// TIA Portal project "EMS" (V15.1)

(* hardware
DEVICE "HMI_SDC"  TP1500 Comfort
   slot 0: "HMI_SDC"  TP1500 Comfort  6AV2 124-0QC02-0AX0  15.0.0.0
   slot 1: "HMI_RT_2"  TP1500 Comfort  6AV2 124-0QC02-0AX0  15.0.0.0
   slot 5: "HMI_SDC._CP_2"  PROFINET Interface  15.0.0.0
      slot 1: "PROFINET Schnittstelle_1"  PROFINET Interface
         slot 1: "Port_1"  Port
         slot 2: "Port_2"  Port
   slot 6: "HMI_SDC._CP_1"  PROFINET Interface  15.0.0.0
      slot 1: "PROFINET Schnittstelle_GBit"  PROFINET Interface
         slot 1: "Port_1"  Port
   slot 7: "HMI_SDC.I/DP_CP_1"  MPI/DP Interface  15.0.0.0
DEVICE "SCALANCE W client"  SCALANCE W-Station
   slot 0: "SCALANCE W rack"  Rail
   slot 0: "_wlan"  SCALANCE W734-1 RJ45 US  6GK5 734-1FX00-0AB0  V6.2
DEVICE "S71500/ET200MP station_1"  S7-1500 station
   slot 0: "Rail_0"  Rack  6ES7 590-1***0-0AA0
   slot 1: "SDC_PLC"  CPU 1518-4 PN/DP  6ES7 518-4AP00-0AB0  V2.6
      slot 3: "CPU display_1"  6ES7591-1BA00-0AA0
   slot 2: "DI 16x24VDC BA_1"  DI 16x24VDC BA  6ES7 521-1BH10-0AA0  V1.0
   slot 3: "DQ 16x24VDC/0.5A BA_1"  DQ 16x24VDC/0.5A BA  6ES7 522-1BH10-0AA0  V1.0
DEVICE "ET 200SP station_2"  ET 200SP-Station
   slot 0: "Rack_0"  Rack  6ES5 710-8MAx1
   slot 1: "_PLC"  CPU 1512SP F-1 PN  6ES7 512-1SK01-0AB0  V2.1
   slot 2: "F-DI 8x24VDC HF_1"  F-DI 8x24VDC HF  6ES7 136-6BA00-0CA0  V1.0
      slot 1: "F-DI 8x24VDC HF_1"  F-DI 8x24VDC HF
   slot 3: "F-DQ 4x24VDC/2A PM HF_1"  F-DQ 4x24VDC/2A PM HF  6ES7 136-6DB00-0CA0  V1.0
      slot 1: "F-DQ 4x24VDC/2A PM HF_1"  F-DQ 4x24VDC/2A PM HF
   slot 4: "DI 16x24VDC ST_1"  DI 16x24VDC ST  6ES7 131-6BH00-0BA0  V1.1
      slot 1: "DI 16x24VDC ST_1"  DI 16x24VDC ST
   slot 5: "DQ 8x24VDC/0.5A ST_1"  DQ 8x24VDC/0.5A ST  6ES7 132-6BF01-0BA0  V0.0
      slot 1: "DQ 8x24VDC/0.5A ST_1"  DQ 8x24VDC/0.5A ST
   slot 6: "Server module_1"  Server module  6ES7 193-6PA00-0AA0  V1.1
      slot 1: "Server module_1"  Server module
   slot 127: "BA 2xRJ45"  BA 2xRJ45  6ES7 193-6AR00-0AA0  V0.0
      slot 32769: "Port_1"  6ES7 193-6AR00-0AA0
      slot 32770: "Port_2"  6ES7 193-6AR00-0AA0
DEVICE "GSD device_4"  GSD.Device.PN
   slot 0: "Rack"  Rack  V1.0
   slot 0: "_DRIVE"  SINAMICS G120D CU240D-2 PN(-F) V4.7  6SL3 544-0FB2x-1Fxx  V4.70
      slot 0: "SINAMICS G120D CU240D-2 PN(-F) V4.7"  SINAMICS G120D CU240D-2 PN(-F) V4.7
      slot 1: "PN-IO"  PN-IO
         slot 1: "Port 1"  Port 1
         slot 2: "Port 2"  Port 2
      slot 1: "Drive_1"  Drive
         slot 0: "Module Access Point"  Module Access Point
   slot 2: "SIEMENS telegram 352, PZD-6/6"  SIEMENS telegram 352, PZD-6/6
DEVICE "GSD device_1"  GSD.Device.PN
   slot 0: "Rack"  Rack  V1.0
   slot 0: "_ENCODER"  PCV-F200-B17-6011 Position Encoder  PXVxx-F200-B17-V1D-6011
      slot 0: "PCV-F200-B17-6011 Position Encoder"  PCV-F200-B17-6011 Position Encoder
      slot 1: "Interface"  Interface
         slot 1: "Port 1"  Port 1
         slot 2: "Port 2"  Port 2
      slot 1: "Configuration_1"  Configuration
         slot 0: "Configuration"  Configuration
   slot 2: "status_1"  status
      slot 0: "status"  status
   slot 3: "x position_1"  x position
      slot 0: "x position"  x position
   slot 4: "y position_1"  y position
      slot 0: "y position"  y position
DEVICE "GSD device_6"  GSD.Device.PN
   slot 0: "Rack"  Rack  V1.0
   slot 0: "_HMI"  IRD400  6ES7 292-0AA50-1AA0  R01.00.00
      slot 0: "IRD400"  IRD400
      slot 1: "PNIO"  PNIO
         slot 1: "Port 1"  Port 1
         slot 2: "Port 2"  Port 2
      slot 1: "IR Remote Control_1"  IR Remote Control
         slot 0: "IR Remote Control"  IR Remote Control
      slot 2: "Display and LED _1"  Display and LED 
         slot 0: "Display and LED"  Display and LED 
      slot 3: "DIO_1"  DIO
         slot 0: "DIO"  DIO
      slot 4: "IR-P2P_1"  IR-P2P
         slot 0: "IR-P2P"  IR-P2P
      slot 5: "Device Control_1"  Device Control
         slot 0: "Device Control"  Device Control
DEVICE "SCALANCE W access point"  SCALANCE W-Station
   slot 0: "SCALANCE W rack"  Rail
   slot 0: "WLAN_1"  SCALANCE W788-1 M12 US  6GK5 788-1GD00-0AB0  V6.2
DEVICE "GSD device_11"  GSD.Device.PN
   slot 0: "Rack"  Rack  V1.0
   slot 0: "plx32-pnd"  PLX32-EIP-PND  EPD2  1.02.002
      slot 0: "PLX32-EIP-PND"  PLX32-EIP-PND
      slot 1: "Interface1"  Interface1
         slot 1: "Port1"  Port1
   slot 1: "INPUT 512 Byte_1"  INPUT 512 Byte
      slot 0: "INPUT 512 Byte"  INPUT 512 Byte
   slot 2: "OUTPUT 512 Byte_1"  OUTPUT 512 Byte
      slot 0: "OUTPUT 512 Byte"  OUTPUT 512 Byte
   slot 3: "INPUT 256 Byte_3"  INPUT 256 Byte
      slot 0: "INPUT 256 Byte"  INPUT 256 Byte
   slot 4: "OUTPUT 256 Byte_3"  OUTPUT 256 Byte
      slot 0: "OUTPUT 256 Byte"  OUTPUT 256 Byte
   slot 5: "INPUT 256 Byte_2"  INPUT 256 Byte
      slot 0: "INPUT 256 Byte"  INPUT 256 Byte
   slot 6: "OUTPUT 256 Byte_2"  OUTPUT 256 Byte
      slot 0: "OUTPUT 256 Byte"  OUTPUT 256 Byte
   slot 7: "INPUT 256 Byte_1"  INPUT 256 Byte
      slot 0: "INPUT 256 Byte"  INPUT 256 Byte
   slot 8: "OUTPUT 256 Byte_1"  OUTPUT 256 Byte
      slot 0: "OUTPUT 256 Byte"  OUTPUT 256 Byte
*)

// ===== PLC "SDC_PLC"  CPU 1518-4 PN/DP =====

VAR_GLOBAL   // PLC tag table "Default tag table"
   "LinePLC1_RD_ready" AT %I4248.0 : Bool;
   "EMS_ProductionSpeedRef" AT %IW6130 : Word;
   "EMS_CarrierSpeedRef" AT %IW6126 : Word;
   "SDC_C2_OUT_W9" AT %QW468 : Word;
   "System_Byte" AT %MB1 : Byte;
   "FirstScan" AT %M1.0 : Bool;
   "DiagStatusUpdate" AT %M1.1 : Bool;
   "AlwaysTRUE" AT %M1.2 : Bool;
   "AlwaysFALSE" AT %M1.3 : Bool;
   "Clock_Byte" AT %MB0 : Byte;
   "Clock_10Hz" AT %M0.0 : Bool;
   "Clock_5Hz" AT %M0.1 : Bool;
   "Clock_2.5Hz" AT %M0.2 : Bool;
   "Clock_2Hz" AT %M0.3 : Bool;
   "Clock_1.25Hz" AT %M0.4 : Bool;
   "Clock_1Hz" AT %M0.5 : Bool;
   "Clock_0.625Hz" AT %M0.6 : Bool;
   "Clock_0.5Hz" AT %M0.7 : Bool;
   "tem" AT %M2.0 : Bool;
   "reset" AT %M2.1 : Bool;
   "ZoneCnt" AT %MW4 : Int;
   "Totalcar" AT %MW6 : Int;
   "Tag_3" AT %M2.2 : Bool;
   "carrierzone" AT %MW8 : Int;
   "Carriercnt" AT %MW10 : Int;
   "Carriercnt(1)" AT %MW12 : Int;
   "carrposn" AT %MW14 : Int;
   "IndexArraytemp" AT %MW20 : Int;
   "tempsort" AT %M2.4 : Bool;
   "tempenable2" AT %M2.5 : Bool;
   "tempenable3" AT %M2.6 : Bool;
   "tempenable4" AT %M2.7 : Bool;
   "tempenable5" AT %M3.0 : Bool;
   "tempenable7" AT %M3.1 : Bool;
   "tempblock" AT %M3.2 : Bool;
   "CarrierCounterGbl" AT %MW16 : Int;
   "temp" AT %M3.3 : Bool;
   "cARRIERTESTPOINT" AT %MW18 : Int;
   "cARRIERTESTPOINTBOOL" AT %M3.4 : Bool;
   "cARIERLOOPCOUNT" AT %MW22 : Int;
   "cARIERLOOPCOUNT2" AT %MW24 : Int;
   "tempcarrier27cmdfwd" AT %MW26 : Int;
   "tempcarrier27cmdfwd1" AT %M3.5 : Bool;
   "ZoneCounterGbl" AT %MW28 : Int;
   "IndiconTempDebugON" AT %M3.6 : Bool;
   "HMI_EMS_Nr" AT %MW30 : Int;
   "HMI_EMS_Nr_Calc1" AT %MW32 : Int;
   "HMI_EMS_Nr_Calc2" AT %MW34 : Int;
   "HMI_EMS_Nr__Flt_Out" AT %MW36 : Int;
   "HMI_EMS_Nr__Warn_Out" AT %MW38 : Int;
   "TrafficCopZoneArrayPosCounter" AT %MW40 : Int;
   "SectionComment" AT %M42.0 : Bool;
   "DuplicateCarrierfound" AT %M42.1 : Bool;
   "FaultReset" AT %M42.2 : Bool;
   "DuplicateCarrierNumber" AT %MW44 : Word;
   "CarrierNumberLoop" AT %MW46 : Int;
   "Zone5_ClearToEnter" AT %M42.3 : Bool;
   "PrevCarrierInTransitMem" AT %M42.4 : Bool;
   "SecondDuplicateCarrierPosition" AT %MW50 : Word;
   "FirstDuplicateCarrierPosition" AT %MW48 : Word;
   "EMS_Fault_Reset" AT %M42.5 : Bool;
   "TCCarrierCounterGbl" AT %MW100 : Int;
   "FC206CarrierLoop" AT %MW52 : Int;
   "FC206PositionLoop" AT %MW54 : Int;
   "CARRIER01_POSITION_SDC_OUT" AT %ID402 : DWord;
   "Temp_Int" AT %MW56 : Int;
   "CARRIER #01   1 STATUS [0].5" AT %M80.5 : Bool;
   "CARRIER #01   CURRENT" AT %MW72 : Int;
   "CARRIER #01   G120D CONTROL WORD.0" AT %M74.0 : Bool;
   "CARRIER #01   G120D CONTROL WORD.1" AT %M74.1 : Bool;
   "CARRIER #01   G120D CONTROL WORD.10" AT %M75.2 : Bool;
   "CARRIER #01   G120D CONTROL WORD.11" AT %M75.3 : Bool;
   "CARRIER #01   G120D CONTROL WORD.12" AT %M75.4 : Bool;
   "CARRIER #01   G120D CONTROL WORD.13" AT %M75.5 : Bool;
   "CARRIER #01   G120D CONTROL WORD.14" AT %M75.6 : Bool;
   "CARRIER #01   G120D CONTROL WORD.15" AT %M75.7 : Bool;
   "CARRIER #01   G120D CONTROL WORD.2" AT %M74.2 : Bool;
   "CARRIER #01   G120D CONTROL WORD.3" AT %M74.3 : Bool;
   "CARRIER #01   G120D CONTROL WORD.4" AT %M74.4 : Bool;
   "CARRIER #01   G120D CONTROL WORD.5" AT %M74.5 : Bool;
   "CARRIER #01   G120D CONTROL WORD.6" AT %M74.6 : Bool;
   "CARRIER #01   G120D CONTROL WORD.7" AT %M74.7 : Bool;
   "CARRIER #01   G120D CONTROL WORD.8" AT %M75.0 : Bool;
   "CARRIER #01   G120D CONTROL WORD.9" AT %M75.1 : Bool;
   "CARRIER #01   G120D STATUS WORD.0" AT %M76.0 : Bool;
   "CARRIER #01   G120D STATUS WORD.1" AT %M76.1 : Bool;
   "CARRIER #01   G120D STATUS WORD.10" AT %M77.2 : Bool;
   "CARRIER #01   G120D STATUS WORD.11" AT %M77.3 : Bool;
   "CARRIER #01   G120D STATUS WORD.12" AT %M77.4 : Bool;
   "CARRIER #01   G120D STATUS WORD.13" AT %M77.5 : Bool;
   "CARRIER #01   G120D STATUS WORD.14" AT %M77.6 : Bool;
   "CARRIER #01   G120D STATUS WORD.15" AT %M77.7 : Bool;
   "CARRIER #01   G120D STATUS WORD.2" AT %M76.2 : Bool;
   "CARRIER #01   G120D STATUS WORD.3" AT %M76.3 : Bool;
   "CARRIER #01   G120D STATUS WORD.4" AT %M76.4 : Bool;
   "CARRIER #01   G120D STATUS WORD.5" AT %M76.5 : Bool;
   "CARRIER #01   G120D STATUS WORD.6" AT %M76.6 : Bool;
   "CARRIER #01   G120D STATUS WORD.7" AT %M76.7 : Bool;
   "CARRIER #01   G120D STATUS WORD.8" AT %M77.0 : Bool;
   "CARRIER #01   G120D STATUS WORD.9" AT %M77.1 : Bool;
   "CARRIER #01   POSITION" AT %MW78 : Int;
   "CARRIER #01 480VPowerOn_MDCB1" AT %M80.0 : Bool;
   "CARRIER #01 CrashDetectSW" AT %M80.1 : Bool;
   "CARRIER #01 DCsupplyOnPSCB2" AT %M80.2 : Bool;
   "CARRIER #01 FaultLight_LH" AT %M80.3 : Bool;
   "CARRIER #01 FaultLight_RH" AT %M80.4 : Bool;
   "CARRIER #01 PB1_ProdHoldLH" AT %M80.6 : Bool;
   "CARRIER #01 PB2_ResetLH" AT %M80.7 : Bool;
   "CARRIER #01 PB3_ProdHoldRH" AT %M81.0 : Bool;
   "CARRIER #01 PB4_ResetRH" AT %M81.1 : Bool;
   "CARRIER #01 RunLight_LH" AT %M81.2 : Bool;
   "CARRIER #01 RunLight_RH" AT %M81.3 : Bool;
   "CARRIER #01 SitopSelectStatus" AT %M81.4 : Bool;
   "CARRIER #01 SpareInput(2_1)" AT %M81.5 : Bool;
   "CARRIER #01 SpareInput(2_2)" AT %M81.6 : Bool;
   "CARRIER #01 SpareInput(2_3)" AT %M81.7 : Bool;
   "CARRIER #01 SpareInput(2_4)" AT %M82.0 : Bool;
   "CARRIER #01 SpareInput(2_5)" AT %M82.1 : Bool;
   "CARRIER #01 SpareInput(2_6)" AT %M82.2 : Bool;
   "CARRIER #01 SpareInput(2_7)" AT %M82.3 : Bool;
   "CARRIER #01 SpareInput(4_1)" AT %M82.4 : Bool;
   "CARRIER #01 SpareInput(4_14)" AT %M82.5 : Bool;
   "CARRIER #01 SpareInput(4_15)" AT %M82.6 : Bool;
   "CARRIER #01 SpareInput(4_16)" AT %M82.7 : Bool;
   "CARRIER #01 SpareInput(4_17)" AT %M83.0 : Bool;
   "CARRIER #01 SpareInput(4_2)" AT %M83.1 : Bool;
   "CARRIER #01 SpareInput(4_5)" AT %M83.2 : Bool;
   "CARRIER #01 SpareInput(4_6)" AT %M83.3 : Bool;
   "CARRIER #01 SpareInput(4_7)" AT %M83.4 : Bool;
   "CARRIER #01 SpareOutput(5_5)" AT %M83.5 : Bool;
   "CARRIER #01 SpareOutput(5_6)" AT %M83.6 : Bool;
   "CARRIER #01 SpareOutput(5_7)" AT %M83.7 : Bool;
   "CARRIER #01 SpareSafetyOutput(3_1)" AT %M84.0 : Bool;
   "CARRIER #01 SpareSafetyOutput(3_2)" AT %M84.1 : Bool;
   "CARRIER #01 SpareSafetyOutput(3_3)" AT %M84.2 : Bool;
   "CARRIER #01 SpareSafetyOutput(3_4)" AT %M84.3 : Bool;
   "CARRIER #01 SpareSafetyOutput(3_5)" AT %M84.4 : Bool;
   "CARRIER #01 SpareSafetyOutput(3_6)" AT %M84.5 : Bool;
   "CARRIER #01 SpareSafetyOutput(3_7)" AT %M84.6 : Bool;
   "Carrier #01_ At Command Position" AT %M84.7 : Bool;
   "Carrier #01_ Carrier in zone" AT %MW86 : Int;
   "Carrier #01_ Next carrier number" AT %MW88 : Int;
   "Carrier 1  Drive Status" AT %I412.1 : Bool;
   "Carrier 1 HMI Status" AT %I412.2 : Bool;
   "Carrier 1 PnF Encoder Status" AT %I412.0 : Bool;
   "Carrier 1 Profinet Fault" AT %I410.7 : Bool;
   "Carrier 2  Drive Status" AT %I432.1 : Bool;
   "Carrier 2 HMI Status" AT %I432.2 : Bool;
   "Carrier 2 PnF Encoder Status" AT %I432.0 : Bool;
   "Carrier 2 Profinet Fault" AT %I430.7 : Bool;
   "Carrier 3  Drive Status" AT %I452.1 : Bool;
   "Carrier 3 HMI Status" AT %I452.2 : Bool;
   "Carrier 3 PnF Encoder Status" AT %I452.0 : Bool;
   "Carrier 4  Drive Status" AT %I472.1 : Bool;
   "Carrier 4 HMI Status" AT %I472.2 : Bool;
   "Carrier 4 PnF Encoder Status" AT %I472.0 : Bool;
   "Carrier 4 Profinet Fault" AT %I470.7 : Bool;
   "Carrier_Index_HMI" AT %MW70 : Int;
   "HMI_Zone_Nr" AT %MW102 : Int;
END_VAR

VAR_GLOBAL CONSTANT   // PLC tag table "UserDiag_Constants"
   "USERDIAG_IOSYSTEM_1" : Int := 1;   // Index for first IO-System/DP-Mastersystem
   "USERDIAG_IOSYSTEM_2" : Int := 2;   // Index for second IO-System/DP-Mastersystem
   "USERDIAG_DEVICES_PER_SCREEN_UPPER_LIM" : Int := 128;   // Upper limit of devices per HMI screen
   "USERDIAG_SLOTS_PER_SCREEN_UPPER_LIM" : Int := 31;   // Upper limit of slots per HMI screen
   "USERDIAG_SLOTS_PER_DEVICE_UPPER_LIM" : Int := 31;   // max number of modules per device
   "USERDIAG_DEVICES_PER_IO_SYSTEM_UPPER_LIM" : Int := 128;   // Upper limit of devices/slaves per IO-System/DP-Mastersystem
   "USERDIAG_SLOTS_PER_PLC_UPPER_LIM" : Int := 31;   // max number of local modules
   "USERDIAG_IO_SYSTEMS_UPPER_LIM" : Int := 2;   // Upper limit of IO-Systems/DP-Mastersystems
   "USERDIAG_IOSYSTEM_3" : Int := 3;   // Index for third IO-System/DP-Mastersystem
END_VAR

VAR_GLOBAL   // PLC tag table "SDC_AB_TagTable"
   "SDC_EMS01_CARRIER1_Spare0" AT %Q6768.0 : Bool;
   "SDC_EMS01_CARRIER1_DriveTripped" AT %Q6768.1 : Bool;
   "SDC_EMS01_CARRIER1_Spare2" AT %Q6768.2 : Bool;
   "SDC_EMS01_CARRIER1_PositioningComplete" AT %Q6768.3 : Bool;
   "SDC_EMS01_CARRIER1_RunStopPressed" AT %Q6768.4 : Bool;
   "SDC_EMS01_CARRIER1_Moving" AT %Q6768.5 : Bool;
   "SDC_EMS01_CARRIER1_Faulted" AT %Q6768.6 : Bool;
   "SDC_EMS01_CARRIER1_InAuto" AT %Q6768.7 : Bool;
   "SDC_EMS01_CARRIER2_Spare0" AT %Q6769.0 : Bool;
   "SDC_EMS01_CARRIER2_DriveTripped" AT %Q6769.1 : Bool;
   "SDC_EMS01_CARRIER2_Spare2" AT %Q6769.2 : Bool;
   "SDC_EMS01_CARRIER2_PositioningComplete" AT %Q6769.3 : Bool;
   "SDC_EMS01_CARRIER2_RunStopPressed" AT %Q6769.4 : Bool;
   "SDC_EMS01_CARRIER2_Moving" AT %Q6769.5 : Bool;
   "SDC_EMS01_CARRIER2_Faulted" AT %Q6769.6 : Bool;
   "SDC_EMS01_CARRIER2_InAuto" AT %Q6769.7 : Bool;
   "SDC_EMS01_CARRIER3_Spare0" AT %Q6770.0 : Bool;
   "SDC_EMS01_CARRIER3_DriveTripped" AT %Q6770.1 : Bool;
   "SDC_EMS01_CARRIER3_Spare2" AT %Q6770.2 : Bool;
   "SDC_EMS01_CARRIER3_PositioningComplete" AT %Q6770.3 : Bool;
   "SDC_EMS01_CARRIER3_RunStopPressed" AT %Q6770.4 : Bool;
   "SDC_EMS01_CARRIER3_Moving" AT %Q6770.5 : Bool;
   "SDC_EMS01_CARRIER3_Faulted" AT %Q6770.6 : Bool;
   "SDC_EMS01_CARRIER3_InAuto" AT %Q6770.7 : Bool;
   "SDC_EMS01_CARRIER4_Spare0" AT %Q6771.0 : Bool;
   "SDC_EMS01_CARRIER4_DriveTripped" AT %Q6771.1 : Bool;
   "SDC_EMS01_CARRIER4_Spare2" AT %Q6771.2 : Bool;
   "SDC_EMS01_CARRIER4_PositioningComplete" AT %Q6771.3 : Bool;
   "SDC_EMS01_CARRIER4_RunStopPressed" AT %Q6771.4 : Bool;
   "SDC_EMS01_CARRIER4_Moving" AT %Q6771.5 : Bool;
   "SDC_EMS01_CARRIER4_Faulted" AT %Q6771.6 : Bool;
   "SDC_EMS01_CARRIER4_InAuto" AT %Q6771.7 : Bool;
   "SDC_EMS01_CARRIER5_Spare0" AT %Q6772.0 : Bool;
   "SDC_EMS01_CARRIER5_DriveTripped" AT %Q6772.1 : Bool;
   "SDC_EMS01_CARRIER5_Spare2" AT %Q6772.2 : Bool;
   "SDC_EMS01_CARRIER5_PositioningComplete" AT %Q6772.3 : Bool;
   "SDC_EMS01_CARRIER5_RunStopPressed" AT %Q6772.4 : Bool;
   "SDC_EMS01_CARRIER5_Moving" AT %Q6772.5 : Bool;
   "SDC_EMS01_CARRIER5_Faulted" AT %Q6772.6 : Bool;
   "SDC_EMS01_CARRIER5_InAuto" AT %Q6772.7 : Bool;
   "SDC_EMS01_CARRIER6_Spare0" AT %Q6773.0 : Bool;
   "SDC_EMS01_CARRIER6_DriveTripped" AT %Q6773.1 : Bool;
   "SDC_EMS01_CARRIER6_Spare2" AT %Q6773.2 : Bool;
   "SDC_EMS01_CARRIER6_PositioningComplete" AT %Q6773.3 : Bool;
   "SDC_EMS01_CARRIER6_RunStopPressed" AT %Q6773.4 : Bool;
   "SDC_EMS01_CARRIER6_Moving" AT %Q6773.5 : Bool;
   "SDC_EMS01_CARRIER6_Faulted" AT %Q6773.6 : Bool;
   "SDC_EMS01_CARRIER6_InAuto" AT %Q6773.7 : Bool;
   "SDC_EMS01_CARRIER7_Spare0" AT %Q6774.0 : Bool;
   "SDC_EMS01_CARRIER7_DriveTripped" AT %Q6774.1 : Bool;
   "SDC_EMS01_CARRIER7_Spare2" AT %Q6774.2 : Bool;
   "SDC_EMS01_CARRIER7_PositioningComplete" AT %Q6774.3 : Bool;
   "SDC_EMS01_CARRIER7_RunStopPressed" AT %Q6774.4 : Bool;
   "SDC_EMS01_CARRIER7_Moving" AT %Q6774.5 : Bool;
   "SDC_EMS01_CARRIER7_Faulted" AT %Q6774.6 : Bool;
   "SDC_EMS01_CARRIER7_InAuto" AT %Q6774.7 : Bool;
   "SDC_EMS01_CARRIER8_Spare0" AT %Q6775.0 : Bool;
   "SDC_EMS01_CARRIER8_DriveTripped" AT %Q6775.1 : Bool;
   "SDC_EMS01_CARRIER8_Spare2" AT %Q6775.2 : Bool;
   "SDC_EMS01_CARRIER8_PositioningComplete" AT %Q6775.3 : Bool;
   "SDC_EMS01_CARRIER8_RunStopPressed" AT %Q6775.4 : Bool;
   "SDC_EMS01_CARRIER8_Moving" AT %Q6775.5 : Bool;
   "SDC_EMS01_CARRIER8_Faulted" AT %Q6775.6 : Bool;
   "SDC_EMS01_CARRIER8_InAuto" AT %Q6775.7 : Bool;
   "SDC_EMS01_CARRIER9_Spare0" AT %Q6776.0 : Bool;
   "SDC_EMS01_CARRIER9_DriveTripped" AT %Q6776.1 : Bool;
   "SDC_EMS01_CARRIER9_Spare2" AT %Q6776.2 : Bool;
   "SDC_EMS01_CARRIER9_PositioningComplete" AT %Q6776.3 : Bool;
   "SDC_EMS01_CARRIER9_RunStopPressed" AT %Q6776.4 : Bool;
   "SDC_EMS01_CARRIER9_Moving" AT %Q6776.5 : Bool;
   "SDC_EMS01_CARRIER9_Faulted" AT %Q6776.6 : Bool;
   "SDC_EMS01_CARRIER9_InAuto" AT %Q6776.7 : Bool;
   "SDC_EMS01_CARRIER10_Spare0" AT %Q6777.0 : Bool;
   "SDC_EMS01_CARRIER10_DriveTripped" AT %Q6777.1 : Bool;
   "SDC_EMS01_CARRIER10_Spare2" AT %Q6777.2 : Bool;
   "SDC_EMS01_CARRIER10_PositioningComplete" AT %Q6777.3 : Bool;
   "SDC_EMS01_CARRIER10_RunStopPressed" AT %Q6777.4 : Bool;
   "SDC_EMS01_CARRIER10_Moving" AT %Q6777.5 : Bool;
   "SDC_EMS01_CARRIER10_Faulted" AT %Q6777.6 : Bool;
   "SDC_EMS01_CARRIER10_InAuto" AT %Q6777.7 : Bool;
   "SDC_EMS01_CARRIER11_Spare0" AT %Q6778.0 : Bool;
   "SDC_EMS01_CARRIER11_DriveTripped" AT %Q6778.1 : Bool;
   "SDC_EMS01_CARRIER11_Spare2" AT %Q6778.2 : Bool;
   "SDC_EMS01_CARRIER11_PositioningComplete" AT %Q6778.3 : Bool;
   "SDC_EMS01_CARRIER11_RunStopPressed" AT %Q6778.4 : Bool;
   "SDC_EMS01_CARRIER11_Moving" AT %Q6778.5 : Bool;
   "SDC_EMS01_CARRIER11_Faulted" AT %Q6778.6 : Bool;
   "SDC_EMS01_CARRIER11_InAuto" AT %Q6778.7 : Bool;
   "SDC_EMS01_CARRIER12_Spare0" AT %Q6779.0 : Bool;
   "SDC_EMS01_CARRIER12_DriveTripped" AT %Q6779.1 : Bool;
   "SDC_EMS01_CARRIER12_Spare2" AT %Q6779.2 : Bool;
   "SDC_EMS01_CARRIER12_PositioningComplete" AT %Q6779.3 : Bool;
   "SDC_EMS01_CARRIER12_RunStopPressed" AT %Q6779.4 : Bool;
   "SDC_EMS01_CARRIER12_Moving" AT %Q6779.5 : Bool;
   "SDC_EMS01_CARRIER12_Faulted" AT %Q6779.6 : Bool;
   "SDC_EMS01_CARRIER12_InAuto" AT %Q6779.7 : Bool;
   "SDC_EMS01_CARRIER13_Spare0" AT %Q6780.0 : Bool;
   "SDC_EMS01_CARRIER13_DriveTripped" AT %Q6780.1 : Bool;
   "SDC_EMS01_CARRIER13_Spare2" AT %Q6780.2 : Bool;
   "SDC_EMS01_CARRIER13_PositioningComplete" AT %Q6780.3 : Bool;
   "SDC_EMS01_CARRIER13_RunStopPressed" AT %Q6780.4 : Bool;
   "SDC_EMS01_CARRIER13_Moving" AT %Q6780.5 : Bool;
   "SDC_EMS01_CARRIER13_Faulted" AT %Q6780.6 : Bool;
   "SDC_EMS01_CARRIER13_InAuto" AT %Q6780.7 : Bool;
   "SDC_EMS01_CARRIER14_Spare0" AT %Q6781.0 : Bool;
   "SDC_EMS01_CARRIER14_DriveTripped" AT %Q6781.1 : Bool;
   "SDC_EMS01_CARRIER14_Spare2" AT %Q6781.2 : Bool;
   "SDC_EMS01_CARRIER14_PositioningComplete" AT %Q6781.3 : Bool;
   "SDC_EMS01_CARRIER14_RunStopPressed" AT %Q6781.4 : Bool;
   "SDC_EMS01_CARRIER14_Moving" AT %Q6781.5 : Bool;
   "SDC_EMS01_CARRIER14_Faulted" AT %Q6781.6 : Bool;
   "SDC_EMS01_CARRIER14_InAuto" AT %Q6781.7 : Bool;
   "SDC_EMS01_CARRIER15_Spare0" AT %Q6782.0 : Bool;
   "SDC_EMS01_CARRIER15_DriveTripped" AT %Q6782.1 : Bool;
   "SDC_EMS01_CARRIER15_Spare2" AT %Q6782.2 : Bool;
   "SDC_EMS01_CARRIER15_PositioningComplete" AT %Q6782.3 : Bool;
   "SDC_EMS01_CARRIER15_RunStopPressed" AT %Q6782.4 : Bool;
   "SDC_EMS01_CARRIER15_Moving" AT %Q6782.5 : Bool;
   "SDC_EMS01_CARRIER15_Faulted" AT %Q6782.6 : Bool;
   "SDC_EMS01_CARRIER15_InAuto" AT %Q6782.7 : Bool;
   "SDC_EMS01_CARRIER16_Spare0" AT %Q6783.0 : Bool;
   "SDC_EMS01_CARRIER16_DriveTripped" AT %Q6783.1 : Bool;
   "SDC_EMS01_CARRIER16_Spare2" AT %Q6783.2 : Bool;
   "SDC_EMS01_CARRIER16_PositioningComplete" AT %Q6783.3 : Bool;
   "SDC_EMS01_CARRIER16_RunStopPressed" AT %Q6783.4 : Bool;
   "SDC_EMS01_CARRIER16_Moving" AT %Q6783.5 : Bool;
   "SDC_EMS01_CARRIER16_Faulted" AT %Q6783.6 : Bool;
   "SDC_EMS01_CARRIER16_InAuto" AT %Q6783.7 : Bool;
   "SDC_EMS01_CARRIER17_Spare0" AT %Q6784.0 : Bool;
   "SDC_EMS01_CARRIER17_DriveTripped" AT %Q6784.1 : Bool;
   "SDC_EMS01_CARRIER17_Spare2" AT %Q6784.2 : Bool;
   "SDC_EMS01_CARRIER17_PositioningComplete" AT %Q6784.3 : Bool;
   "SDC_EMS01_CARRIER17_RunStopPressed" AT %Q6784.4 : Bool;
   "SDC_EMS01_CARRIER17_Moving" AT %Q6784.5 : Bool;
   "SDC_EMS01_CARRIER17_Faulted" AT %Q6784.6 : Bool;
   "SDC_EMS01_CARRIER17_InAuto" AT %Q6784.7 : Bool;
   "SDC_EMS01_CARRIER18_Spare0" AT %Q6785.0 : Bool;
   "SDC_EMS01_CARRIER18_DriveTripped" AT %Q6785.1 : Bool;
   "SDC_EMS01_CARRIER18_Spare2" AT %Q6785.2 : Bool;
   "SDC_EMS01_CARRIER18_PositioningComplete" AT %Q6785.3 : Bool;
   "SDC_EMS01_CARRIER18_RunStopPressed" AT %Q6785.4 : Bool;
   "SDC_EMS01_CARRIER18_Moving" AT %Q6785.5 : Bool;
   "SDC_EMS01_CARRIER18_Faulted" AT %Q6785.6 : Bool;
   "SDC_EMS01_CARRIER18_InAuto" AT %Q6785.7 : Bool;
   "SDC_EMS01_CARRIER19_Spare0" AT %Q6786.0 : Bool;
   "SDC_EMS01_CARRIER19_DriveTripped" AT %Q6786.1 : Bool;
   "SDC_EMS01_CARRIER19_Spare2" AT %Q6786.2 : Bool;
   "SDC_EMS01_CARRIER19_PositioningComplete" AT %Q6786.3 : Bool;
   "SDC_EMS01_CARRIER19_RunStopPressed" AT %Q6786.4 : Bool;
   "SDC_EMS01_CARRIER19_Moving" AT %Q6786.5 : Bool;
   "SDC_EMS01_CARRIER19_Faulted" AT %Q6786.6 : Bool;
   "SDC_EMS01_CARRIER19_InAuto" AT %Q6786.7 : Bool;
   "SDC_EMS01_CARRIER20_Spare0" AT %Q6787.0 : Bool;
   "SDC_EMS01_CARRIER20_DriveTripped" AT %Q6787.1 : Bool;
   "SDC_EMS01_CARRIER20_Spare2" AT %Q6787.2 : Bool;
   "SDC_EMS01_CARRIER20_PositioningComplete" AT %Q6787.3 : Bool;
   "SDC_EMS01_CARRIER20_RunStopPressed" AT %Q6787.4 : Bool;
   "SDC_EMS01_CARRIER20_Moving" AT %Q6787.5 : Bool;
   "SDC_EMS01_CARRIER20_Faulted" AT %Q6787.6 : Bool;
   "SDC_EMS01_CARRIER20_InAuto" AT %Q6787.7 : Bool;
   "SDC_EMS01_CARRIER21_Spare0" AT %Q6788.0 : Bool;
   "SDC_EMS01_CARRIER21_DriveTripped" AT %Q6788.1 : Bool;
   "SDC_EMS01_CARRIER21_Spare2" AT %Q6788.2 : Bool;
   "SDC_EMS01_CARRIER21_PositioningComplete" AT %Q6788.3 : Bool;
   "SDC_EMS01_CARRIER21_RunStopPressed" AT %Q6788.4 : Bool;
   "SDC_EMS01_CARRIER21_Moving" AT %Q6788.5 : Bool;
   "SDC_EMS01_CARRIER21_Faulted" AT %Q6788.6 : Bool;
   "SDC_EMS01_CARRIER21_InAuto" AT %Q6788.7 : Bool;
   "SDC_EMS01_CARRIER22_Spare0" AT %Q6789.0 : Bool;
   "SDC_EMS01_CARRIER22_DriveTripped" AT %Q6789.1 : Bool;
   "SDC_EMS01_CARRIER22_Spare2" AT %Q6789.2 : Bool;
   "SDC_EMS01_CARRIER22_PositioningComplete" AT %Q6789.3 : Bool;
   "SDC_EMS01_CARRIER22_RunStopPressed" AT %Q6789.4 : Bool;
   "SDC_EMS01_CARRIER22_Moving" AT %Q6789.5 : Bool;
   "SDC_EMS01_CARRIER22_Faulted" AT %Q6789.6 : Bool;
   "SDC_EMS01_CARRIER22_InAuto" AT %Q6789.7 : Bool;
   "SDC_EMS01_CARRIER23_Spare0" AT %Q6790.0 : Bool;
   "SDC_EMS01_CARRIER23_DriveTripped" AT %Q6790.1 : Bool;
   "SDC_EMS01_CARRIER23_Spare2" AT %Q6790.2 : Bool;
   "SDC_EMS01_CARRIER23_PositioningComplete" AT %Q6790.3 : Bool;
   "SDC_EMS01_CARRIER23_RunStopPressed" AT %Q6790.4 : Bool;
   "SDC_EMS01_CARRIER23_Moving" AT %Q6790.5 : Bool;
   "SDC_EMS01_CARRIER23_Faulted" AT %Q6790.6 : Bool;
   "SDC_EMS01_CARRIER23_InAuto" AT %Q6790.7 : Bool;
   "SDC_EMS01_CARRIER24_Spare0" AT %Q6791.0 : Bool;
   "SDC_EMS01_CARRIER24_DriveTripped" AT %Q6791.1 : Bool;
   "SDC_EMS01_CARRIER24_Spare2" AT %Q6791.2 : Bool;
   "SDC_EMS01_CARRIER24_PositioningComplete" AT %Q6791.3 : Bool;
   "SDC_EMS01_CARRIER24_RunStopPressed" AT %Q6791.4 : Bool;
   "SDC_EMS01_CARRIER24_Moving" AT %Q6791.5 : Bool;
   "SDC_EMS01_CARRIER24_Faulted" AT %Q6791.6 : Bool;
   "SDC_EMS01_CARRIER24_InAuto" AT %Q6791.7 : Bool;
   "SDC_EMS01_CARRIER25_Spare0" AT %Q6792.0 : Bool;
   "SDC_EMS01_CARRIER25_DriveTripped" AT %Q6792.1 : Bool;
   "SDC_EMS01_CARRIER25_Spare2" AT %Q6792.2 : Bool;
   "SDC_EMS01_CARRIER25_PositioningComplete" AT %Q6792.3 : Bool;
   "SDC_EMS01_CARRIER25_RunStopPressed" AT %Q6792.4 : Bool;
   "SDC_EMS01_CARRIER25_Moving" AT %Q6792.5 : Bool;
   "SDC_EMS01_CARRIER25_Faulted" AT %Q6792.6 : Bool;
   "SDC_EMS01_CARRIER25_InAuto" AT %Q6792.7 : Bool;
   "SDC_EMS01_CARRIER26_Spare0" AT %Q6793.0 : Bool;
   "SDC_EMS01_CARRIER26_DriveTripped" AT %Q6793.1 : Bool;
   "SDC_EMS01_CARRIER26_Spare2" AT %Q6793.2 : Bool;
   "SDC_EMS01_CARRIER26_PositioningComplete" AT %Q6793.3 : Bool;
   "SDC_EMS01_CARRIER26_RunStopPressed" AT %Q6793.4 : Bool;
   "SDC_EMS01_CARRIER26_Moving" AT %Q6793.5 : Bool;
   "SDC_EMS01_CARRIER26_Faulted" AT %Q6793.6 : Bool;
   "SDC_EMS01_CARRIER26_InAuto" AT %Q6793.7 : Bool;
   "SDC_EMS01_CARRIER27_Spare0" AT %Q6794.0 : Bool;
   "SDC_EMS01_CARRIER27_DriveTripped" AT %Q6794.1 : Bool;
   "SDC_EMS01_CARRIER27_Spare2" AT %Q6794.2 : Bool;
   "SDC_EMS01_CARRIER27_PositioningComplete" AT %Q6794.3 : Bool;
   "SDC_EMS01_CARRIER27_RunStopPressed" AT %Q6794.4 : Bool;
   "SDC_EMS01_CARRIER27_Moving" AT %Q6794.5 : Bool;
   "SDC_EMS01_CARRIER27_Faulted" AT %Q6794.6 : Bool;
   "SDC_EMS01_CARRIER27_InAuto" AT %Q6794.7 : Bool;
   "SDC_EMS01_CARRIER28_Spare0" AT %Q6795.0 : Bool;
   "SDC_EMS01_CARRIER28_DriveTripped" AT %Q6795.1 : Bool;
   "SDC_EMS01_CARRIER28_Spare2" AT %Q6795.2 : Bool;
   "SDC_EMS01_CARRIER28_PositioningComplete" AT %Q6795.3 : Bool;
   "SDC_EMS01_CARRIER28_RunStopPressed" AT %Q6795.4 : Bool;
   "SDC_EMS01_CARRIER28_Moving" AT %Q6795.5 : Bool;
   "SDC_EMS01_CARRIER28_Faulted" AT %Q6795.6 : Bool;
   "SDC_EMS01_CARRIER28_InAuto" AT %Q6795.7 : Bool;
   "SDC_EMS01_CARRIER29_Spare0" AT %Q6796.0 : Bool;
   "SDC_EMS01_CARRIER29_DriveTripped" AT %Q6796.1 : Bool;
   "SDC_EMS01_CARRIER29_Spare2" AT %Q6796.2 : Bool;
   "SDC_EMS01_CARRIER29_PositioningComplete" AT %Q6796.3 : Bool;
   "SDC_EMS01_CARRIER29_RunStopPressed" AT %Q6796.4 : Bool;
   "SDC_EMS01_CARRIER29_Moving" AT %Q6796.5 : Bool;
   "SDC_EMS01_CARRIER29_Faulted" AT %Q6796.6 : Bool;
   "SDC_EMS01_CARRIER29_InAuto" AT %Q6796.7 : Bool;
   "SDC_EMS01_CARRIER30_Spare0" AT %Q6797.0 : Bool;
   "SDC_EMS01_CARRIER30_DriveTripped" AT %Q6797.1 : Bool;
   "SDC_EMS01_CARRIER30_Spare2" AT %Q6797.2 : Bool;
   "SDC_EMS01_CARRIER30_PositioningComplete" AT %Q6797.3 : Bool;
   "SDC_EMS01_CARRIER30_RunStopPressed" AT %Q6797.4 : Bool;
   "SDC_EMS01_CARRIER30_Moving" AT %Q6797.5 : Bool;
   "SDC_EMS01_CARRIER30_Faulted" AT %Q6797.6 : Bool;
   "SDC_EMS01_CARRIER30_InAuto" AT %Q6797.7 : Bool;
   "SDC_EMS01_CARRIER31_Spare0" AT %Q6798.0 : Bool;
   "SDC_EMS01_CARRIER31_DriveTripped" AT %Q6798.1 : Bool;
   "SDC_EMS01_CARRIER31_Spare2" AT %Q6798.2 : Bool;
   "SDC_EMS01_CARRIER31_PositioningComplete" AT %Q6798.3 : Bool;
   "SDC_EMS01_CARRIER31_RunStopPressed" AT %Q6798.4 : Bool;
   "SDC_EMS01_CARRIER31_Moving" AT %Q6798.5 : Bool;
   "SDC_EMS01_CARRIER31_Faulted" AT %Q6798.6 : Bool;
   "SDC_EMS01_CARRIER31_InAuto" AT %Q6798.7 : Bool;
   "SDC_EMS01_CARRIER32_Spare0" AT %Q6799.0 : Bool;
   "SDC_EMS01_CARRIER32_DriveTripped" AT %Q6799.1 : Bool;
   "SDC_EMS01_CARRIER32_Spare2" AT %Q6799.2 : Bool;
   "SDC_EMS01_CARRIER32_PositioningComplete" AT %Q6799.3 : Bool;
   "SDC_EMS01_CARRIER32_RunStopPressed" AT %Q6799.4 : Bool;
   "SDC_EMS01_CARRIER32_Moving" AT %Q6799.5 : Bool;
   "SDC_EMS01_CARRIER32_Faulted" AT %Q6799.6 : Bool;
   "SDC_EMS01_CARRIER32_InAuto" AT %Q6799.7 : Bool;
   "SDC_EMS01_CARRIER33_Spare0" AT %Q6800.0 : Bool;
   "SDC_EMS01_CARRIER33_DriveTripped" AT %Q6800.1 : Bool;
   "SDC_EMS01_CARRIER33_Spare2" AT %Q6800.2 : Bool;
   "SDC_EMS01_CARRIER33_PositioningComplete" AT %Q6800.3 : Bool;
   "SDC_EMS01_CARRIER33_RunStopPressed" AT %Q6800.4 : Bool;
   "SDC_EMS01_CARRIER33_Moving" AT %Q6800.5 : Bool;
   "SDC_EMS01_CARRIER33_Faulted" AT %Q6800.6 : Bool;
   "SDC_EMS01_CARRIER33_InAuto" AT %Q6800.7 : Bool;
   "SDC_EMS01_CARRIER34_Spare0" AT %Q6801.0 : Bool;
   "SDC_EMS01_CARRIER34_DriveTripped" AT %Q6801.1 : Bool;
   "SDC_EMS01_CARRIER34_Spare2" AT %Q6801.2 : Bool;
   "SDC_EMS01_CARRIER34_PositioningComplete" AT %Q6801.3 : Bool;
   "SDC_EMS01_CARRIER34_RunStopPressed" AT %Q6801.4 : Bool;
   "SDC_EMS01_CARRIER34_Moving" AT %Q6801.5 : Bool;
   "SDC_EMS01_CARRIER34_Faulted" AT %Q6801.6 : Bool;
   "SDC_EMS01_CARRIER34_InAuto" AT %Q6801.7 : Bool;
   "SDC_EMS01_CARRIER35_Spare0" AT %Q6802.0 : Bool;
   "SDC_EMS01_CARRIER35_DriveTripped" AT %Q6802.1 : Bool;
   "SDC_EMS01_CARRIER35_Spare2" AT %Q6802.2 : Bool;
   "SDC_EMS01_CARRIER35_PositioningComplete" AT %Q6802.3 : Bool;
   "SDC_EMS01_CARRIER35_RunStopPressed" AT %Q6802.4 : Bool;
   "SDC_EMS01_CARRIER35_Moving" AT %Q6802.5 : Bool;
   "SDC_EMS01_CARRIER35_Faulted" AT %Q6802.6 : Bool;
   "SDC_EMS01_CARRIER35_InAuto" AT %Q6802.7 : Bool;
   "SDC_EMS01_CARRIER36_Spare0" AT %Q6803.0 : Bool;
   "SDC_EMS01_CARRIER36_DriveTripped" AT %Q6803.1 : Bool;
   "SDC_EMS01_CARRIER36_Spare2" AT %Q6803.2 : Bool;
   "SDC_EMS01_CARRIER36_PositioningComplete" AT %Q6803.3 : Bool;
   "SDC_EMS01_CARRIER36_RunStopPressed" AT %Q6803.4 : Bool;
   "SDC_EMS01_CARRIER36_Moving" AT %Q6803.5 : Bool;
   "SDC_EMS01_CARRIER36_Faulted" AT %Q6803.6 : Bool;
   "SDC_EMS01_CARRIER36_InAuto" AT %Q6803.7 : Bool;
   "SDC_EMS01_CARRIER37_Spare0" AT %Q6804.0 : Bool;
   "SDC_EMS01_CARRIER37_DriveTripped" AT %Q6804.1 : Bool;
   "SDC_EMS01_CARRIER37_Spare2" AT %Q6804.2 : Bool;
   "SDC_EMS01_CARRIER37_PositioningComplete" AT %Q6804.3 : Bool;
   "SDC_EMS01_CARRIER37_RunStopPressed" AT %Q6804.4 : Bool;
   "SDC_EMS01_CARRIER37_Moving" AT %Q6804.5 : Bool;
   "SDC_EMS01_CARRIER37_Faulted" AT %Q6804.6 : Bool;
   "SDC_EMS01_CARRIER37_InAuto" AT %Q6804.7 : Bool;
   "SDC_EMS01_CARRIER38_Spare0" AT %Q6805.0 : Bool;
   "SDC_EMS01_CARRIER38_DriveTripped" AT %Q6805.1 : Bool;
   "SDC_EMS01_CARRIER38_Spare2" AT %Q6805.2 : Bool;
   "SDC_EMS01_CARRIER38_PositioningComplete" AT %Q6805.3 : Bool;
   "SDC_EMS01_CARRIER38_RunStopPressed" AT %Q6805.4 : Bool;
   "SDC_EMS01_CARRIER38_Moving" AT %Q6805.5 : Bool;
   "SDC_EMS01_CARRIER38_Faulted" AT %Q6805.6 : Bool;
   "SDC_EMS01_CARRIER38_InAuto" AT %Q6805.7 : Bool;
   "SDC_EMS01_CARRIER39_Spare0" AT %Q6806.0 : Bool;
   "SDC_EMS01_CARRIER39_DriveTripped" AT %Q6806.1 : Bool;
   "SDC_EMS01_CARRIER39_Spare2" AT %Q6806.2 : Bool;
   "SDC_EMS01_CARRIER39_PositioningComplete" AT %Q6806.3 : Bool;
   "SDC_EMS01_CARRIER39_RunStopPressed" AT %Q6806.4 : Bool;
   "SDC_EMS01_CARRIER39_Moving" AT %Q6806.5 : Bool;
   "SDC_EMS01_CARRIER39_Faulted" AT %Q6806.6 : Bool;
   "SDC_EMS01_CARRIER39_InAuto" AT %Q6806.7 : Bool;
   "SDC_EMS01_CARRIER40_Spare0" AT %Q6807.0 : Bool;
   "SDC_EMS01_CARRIER40_DriveTripped" AT %Q6807.1 : Bool;
   "SDC_EMS01_CARRIER40_Spare2" AT %Q6807.2 : Bool;
   "SDC_EMS01_CARRIER40_PositioningComplete" AT %Q6807.3 : Bool;
   "SDC_EMS01_CARRIER40_RunStopPressed" AT %Q6807.4 : Bool;
   "SDC_EMS01_CARRIER40_Moving" AT %Q6807.5 : Bool;
   "SDC_EMS01_CARRIER40_Faulted" AT %Q6807.6 : Bool;
   "SDC_EMS01_CARRIER40_InAuto" AT %Q6807.7 : Bool;
   "SDC_EMS01_CARRIER41_Spare0" AT %Q6808.0 : Bool;
   "SDC_EMS01_CARRIER41_DriveTripped" AT %Q6808.1 : Bool;
   "SDC_EMS01_CARRIER41_Spare2" AT %Q6808.2 : Bool;
   "SDC_EMS01_CARRIER41_PositioningComplete" AT %Q6808.3 : Bool;
   "SDC_EMS01_CARRIER41_RunStopPressed" AT %Q6808.4 : Bool;
   "SDC_EMS01_CARRIER41_Moving" AT %Q6808.5 : Bool;
   "SDC_EMS01_CARRIER41_Faulted" AT %Q6808.6 : Bool;
   "SDC_EMS01_CARRIER41_InAuto" AT %Q6808.7 : Bool;
   "SDC_EMS01_CARRIER42_Spare0" AT %Q6809.0 : Bool;
   "SDC_EMS01_CARRIER42_DriveTripped" AT %Q6809.1 : Bool;
   "SDC_EMS01_CARRIER42_Spare2" AT %Q6809.2 : Bool;
   "SDC_EMS01_CARRIER42_PositioningComplete" AT %Q6809.3 : Bool;
   "SDC_EMS01_CARRIER42_RunStopPressed" AT %Q6809.4 : Bool;
   "SDC_EMS01_CARRIER42_Moving" AT %Q6809.5 : Bool;
   "SDC_EMS01_CARRIER42_Faulted" AT %Q6809.6 : Bool;
   "SDC_EMS01_CARRIER42_InAuto" AT %Q6809.7 : Bool;
   "SDC_EMS01_CARRIER43_Spare0" AT %Q6810.0 : Bool;
   "SDC_EMS01_CARRIER43_DriveTripped" AT %Q6810.1 : Bool;
   "SDC_EMS01_CARRIER43_Spare2" AT %Q6810.2 : Bool;
   "SDC_EMS01_CARRIER43_PositioningComplete" AT %Q6810.3 : Bool;
   "SDC_EMS01_CARRIER43_RunStopPressed" AT %Q6810.4 : Bool;
   "SDC_EMS01_CARRIER43_Moving" AT %Q6810.5 : Bool;
   "SDC_EMS01_CARRIER43_Faulted" AT %Q6810.6 : Bool;
   "SDC_EMS01_CARRIER43_InAuto" AT %Q6810.7 : Bool;
   "SDC_EMS01_CARRIER44_Spare0" AT %Q6811.0 : Bool;
   "SDC_EMS01_CARRIER44_DriveTripped" AT %Q6811.1 : Bool;
   "SDC_EMS01_CARRIER44_Spare2" AT %Q6811.2 : Bool;
   "SDC_EMS01_CARRIER44_PositioningComplete" AT %Q6811.3 : Bool;
   "SDC_EMS01_CARRIER44_RunStopPressed" AT %Q6811.4 : Bool;
   "SDC_EMS01_CARRIER44_Moving" AT %Q6811.5 : Bool;
   "SDC_EMS01_CARRIER44_Faulted" AT %Q6811.6 : Bool;
   "SDC_EMS01_CARRIER44_InAuto" AT %Q6811.7 : Bool;
   "SDC_EMS01_CARRIER45_Spare0" AT %Q6812.0 : Bool;
   "SDC_EMS01_CARRIER45_DriveTripped" AT %Q6812.1 : Bool;
   "SDC_EMS01_CARRIER45_Spare2" AT %Q6812.2 : Bool;
   "SDC_EMS01_CARRIER45_PositioningComplete" AT %Q6812.3 : Bool;
   "SDC_EMS01_CARRIER45_RunStopPressed" AT %Q6812.4 : Bool;
   "SDC_EMS01_CARRIER45_Moving" AT %Q6812.5 : Bool;
   "SDC_EMS01_CARRIER45_Faulted" AT %Q6812.6 : Bool;
   "SDC_EMS01_CARRIER45_InAuto" AT %Q6812.7 : Bool;
   "SDC_EMS01_CARRIER46_Spare0" AT %Q6813.0 : Bool;
   "SDC_EMS01_CARRIER46_DriveTripped" AT %Q6813.1 : Bool;
   "SDC_EMS01_CARRIER46_Spare2" AT %Q6813.2 : Bool;
   "SDC_EMS01_CARRIER46_PositioningComplete" AT %Q6813.3 : Bool;
   "SDC_EMS01_CARRIER46_RunStopPressed" AT %Q6813.4 : Bool;
   "SDC_EMS01_CARRIER46_Moving" AT %Q6813.5 : Bool;
   "SDC_EMS01_CARRIER46_Faulted" AT %Q6813.6 : Bool;
   "SDC_EMS01_CARRIER46_InAuto" AT %Q6813.7 : Bool;
   "SDC_EMS01_CARRIER47_Spare0" AT %Q6814.0 : Bool;
   "SDC_EMS01_CARRIER47_DriveTripped" AT %Q6814.1 : Bool;
   "SDC_EMS01_CARRIER47_Spare2" AT %Q6814.2 : Bool;
   "SDC_EMS01_CARRIER47_PositioningComplete" AT %Q6814.3 : Bool;
   "SDC_EMS01_CARRIER47_RunStopPressed" AT %Q6814.4 : Bool;
   "SDC_EMS01_CARRIER47_Moving" AT %Q6814.5 : Bool;
   "SDC_EMS01_CARRIER47_Faulted" AT %Q6814.6 : Bool;
   "SDC_EMS01_CARRIER47_InAuto" AT %Q6814.7 : Bool;
   "SDC_EMS01_CARRIER48_Spare0" AT %Q6815.0 : Bool;
   "SDC_EMS01_CARRIER48_DriveTripped" AT %Q6815.1 : Bool;
   "SDC_EMS01_CARRIER48_Spare2" AT %Q6815.2 : Bool;
   "SDC_EMS01_CARRIER48_PositioningComplete" AT %Q6815.3 : Bool;
   "SDC_EMS01_CARRIER48_RunStopPressed" AT %Q6815.4 : Bool;
   "SDC_EMS01_CARRIER48_Moving" AT %Q6815.5 : Bool;
   "SDC_EMS01_CARRIER48_Faulted" AT %Q6815.6 : Bool;
   "SDC_EMS01_CARRIER48_InAuto" AT %Q6815.7 : Bool;
   "SDC_EMS01_CARRIER49_Spare0" AT %Q6816.0 : Bool;
   "SDC_EMS01_CARRIER49_DriveTripped" AT %Q6816.1 : Bool;
   "SDC_EMS01_CARRIER49_Spare2" AT %Q6816.2 : Bool;
   "SDC_EMS01_CARRIER49_PositioningComplete" AT %Q6816.3 : Bool;
   "SDC_EMS01_CARRIER49_RunStopPressed" AT %Q6816.4 : Bool;
   "SDC_EMS01_CARRIER49_Moving" AT %Q6816.5 : Bool;
   "SDC_EMS01_CARRIER49_Faulted" AT %Q6816.6 : Bool;
   "SDC_EMS01_CARRIER49_InAuto" AT %Q6816.7 : Bool;
   "SDC_EMS01_CARRIER50_Spare0" AT %Q6817.0 : Bool;
   "SDC_EMS01_CARRIER50_DriveTripped" AT %Q6817.1 : Bool;
   "SDC_EMS01_CARRIER50_Spare2" AT %Q6817.2 : Bool;
   "SDC_EMS01_CARRIER50_PositioningComplete" AT %Q6817.3 : Bool;
   "SDC_EMS01_CARRIER50_RunStopPressed" AT %Q6817.4 : Bool;
   "SDC_EMS01_CARRIER50_Moving" AT %Q6817.5 : Bool;
   "SDC_EMS01_CARRIER50_Faulted" AT %Q6817.6 : Bool;
   "SDC_EMS01_CARRIER50_InAuto" AT %Q6817.7 : Bool;
   "SDC_EMS01_CARRIER51_Spare0" AT %Q6818.0 : Bool;
   "SDC_EMS01_CARRIER51_DriveTripped" AT %Q6818.1 : Bool;
   "SDC_EMS01_CARRIER51_Spare2" AT %Q6818.2 : Bool;
   "SDC_EMS01_CARRIER51_PositioningComplete" AT %Q6818.3 : Bool;
   "SDC_EMS01_CARRIER51_RunStopPressed" AT %Q6818.4 : Bool;
   "SDC_EMS01_CARRIER51_Moving" AT %Q6818.5 : Bool;
   "SDC_EMS01_CARRIER51_Faulted" AT %Q6818.6 : Bool;
   "SDC_EMS01_CARRIER51_InAuto" AT %Q6818.7 : Bool;
   "SDC_EMS01_CARRIER52_Spare0" AT %Q6819.0 : Bool;
   "SDC_EMS01_CARRIER52_DriveTripped" AT %Q6819.1 : Bool;
   "SDC_EMS01_CARRIER52_Spare2" AT %Q6819.2 : Bool;
   "SDC_EMS01_CARRIER52_PositioningComplete" AT %Q6819.3 : Bool;
   "SDC_EMS01_CARRIER52_RunStopPressed" AT %Q6819.4 : Bool;
   "SDC_EMS01_CARRIER52_Moving" AT %Q6819.5 : Bool;
   "SDC_EMS01_CARRIER52_Faulted" AT %Q6819.6 : Bool;
   "SDC_EMS01_CARRIER52_InAuto" AT %Q6819.7 : Bool;
   "SDC_EMS01_CARRIER53_Spare0" AT %Q6820.0 : Bool;
   "SDC_EMS01_CARRIER53_DriveTripped" AT %Q6820.1 : Bool;
   "SDC_EMS01_CARRIER53_Spare2" AT %Q6820.2 : Bool;
   "SDC_EMS01_CARRIER53_PositioningComplete" AT %Q6820.3 : Bool;
   "SDC_EMS01_CARRIER53_RunStopPressed" AT %Q6820.4 : Bool;
   "SDC_EMS01_CARRIER53_Moving" AT %Q6820.5 : Bool;
   "SDC_EMS01_CARRIER53_Faulted" AT %Q6820.6 : Bool;
   "SDC_EMS01_CARRIER53_InAuto" AT %Q6820.7 : Bool;
   "SDC_EMS01_CARRIER54_Spare0" AT %Q6821.0 : Bool;
   "SDC_EMS01_CARRIER54_DriveTripped" AT %Q6821.1 : Bool;
   "SDC_EMS01_CARRIER54_Spare2" AT %Q6821.2 : Bool;
   "SDC_EMS01_CARRIER54_PositioningComplete" AT %Q6821.3 : Bool;
   "SDC_EMS01_CARRIER54_RunStopPressed" AT %Q6821.4 : Bool;
   "SDC_EMS01_CARRIER54_Moving" AT %Q6821.5 : Bool;
   "SDC_EMS01_CARRIER54_Faulted" AT %Q6821.6 : Bool;
   "SDC_EMS01_CARRIER54_InAuto" AT %Q6821.7 : Bool;
   "SDC_EMS01_CARRIER55_Spare0" AT %Q6822.0 : Bool;
   "SDC_EMS01_CARRIER55_DriveTripped" AT %Q6822.1 : Bool;
   "SDC_EMS01_CARRIER55_Spare2" AT %Q6822.2 : Bool;
   "SDC_EMS01_CARRIER55_PositioningComplete" AT %Q6822.3 : Bool;
   "SDC_EMS01_CARRIER55_RunStopPressed" AT %Q6822.4 : Bool;
   "SDC_EMS01_CARRIER55_Moving" AT %Q6822.5 : Bool;
   "SDC_EMS01_CARRIER55_Faulted" AT %Q6822.6 : Bool;
   "SDC_EMS01_CARRIER55_InAuto" AT %Q6822.7 : Bool;
   "SDC_EMS01_CARRIER56_Spare0" AT %Q6823.0 : Bool;
   "SDC_EMS01_CARRIER56_DriveTripped" AT %Q6823.1 : Bool;
   "SDC_EMS01_CARRIER56_Spare2" AT %Q6823.2 : Bool;
   "SDC_EMS01_CARRIER56_PositioningComplete" AT %Q6823.3 : Bool;
   "SDC_EMS01_CARRIER56_RunStopPressed" AT %Q6823.4 : Bool;
   "SDC_EMS01_CARRIER56_Moving" AT %Q6823.5 : Bool;
   "SDC_EMS01_CARRIER56_Faulted" AT %Q6823.6 : Bool;
   "SDC_EMS01_CARRIER56_InAuto" AT %Q6823.7 : Bool;
   "SDC_EMS01_CARRIER57_Spare0" AT %Q6824.0 : Bool;
   "SDC_EMS01_CARRIER57_DriveTripped" AT %Q6824.1 : Bool;
   "SDC_EMS01_CARRIER57_Spare2" AT %Q6824.2 : Bool;
   "SDC_EMS01_CARRIER57_PositioningComplete" AT %Q6824.3 : Bool;
   "SDC_EMS01_CARRIER57_RunStopPressed" AT %Q6824.4 : Bool;
   "SDC_EMS01_CARRIER57_Moving" AT %Q6824.5 : Bool;
   "SDC_EMS01_CARRIER57_Faulted" AT %Q6824.6 : Bool;
   "SDC_EMS01_CARRIER57_InAuto" AT %Q6824.7 : Bool;
   "SDC_EMS01_CARRIER58_Spare0" AT %Q6825.0 : Bool;
   "SDC_EMS01_CARRIER58_DriveTripped" AT %Q6825.1 : Bool;
   "SDC_EMS01_CARRIER58_Spare2" AT %Q6825.2 : Bool;
   "SDC_EMS01_CARRIER58_PositioningComplete" AT %Q6825.3 : Bool;
   "SDC_EMS01_CARRIER58_RunStopPressed" AT %Q6825.4 : Bool;
   "SDC_EMS01_CARRIER58_Moving" AT %Q6825.5 : Bool;
   "SDC_EMS01_CARRIER58_Faulted" AT %Q6825.6 : Bool;
   "SDC_EMS01_CARRIER58_InAuto" AT %Q6825.7 : Bool;
   "SDC_EMS01_CARRIER59_Spare0" AT %Q6826.0 : Bool;
   "SDC_EMS01_CARRIER59_DriveTripped" AT %Q6826.1 : Bool;
   "SDC_EMS01_CARRIER59_Spare2" AT %Q6826.2 : Bool;
   "SDC_EMS01_CARRIER59_PositioningComplete" AT %Q6826.3 : Bool;
   "SDC_EMS01_CARRIER59_RunStopPressed" AT %Q6826.4 : Bool;
   "SDC_EMS01_CARRIER59_Moving" AT %Q6826.5 : Bool;
   "SDC_EMS01_CARRIER59_Faulted" AT %Q6826.6 : Bool;
   "SDC_EMS01_CARRIER59_InAuto" AT %Q6826.7 : Bool;
   "SDC_EMS01_CARRIER60_Spare0" AT %Q6827.0 : Bool;
   "SDC_EMS01_CARRIER60_DriveTripped" AT %Q6827.1 : Bool;
   "SDC_EMS01_CARRIER60_Spare2" AT %Q6827.2 : Bool;
   "SDC_EMS01_CARRIER60_PositioningComplete" AT %Q6827.3 : Bool;
   "SDC_EMS01_CARRIER60_RunStopPressed" AT %Q6827.4 : Bool;
   "SDC_EMS01_CARRIER60_Moving" AT %Q6827.5 : Bool;
   "SDC_EMS01_CARRIER60_Faulted" AT %Q6827.6 : Bool;
   "SDC_EMS01_CARRIER60_InAuto" AT %Q6827.7 : Bool;
   "SDC_EMS01_CARRIER61_Spare0" AT %Q6828.0 : Bool;
   "SDC_EMS01_CARRIER61_DriveTripped" AT %Q6828.1 : Bool;